   //-----------------------------
   // HP indication mixinghead 01:
   //-----------------------------
         A     "DB619_State_MPart".Recirculation[1].Lamp_HP."01";
         =     "DB123_MH_IO_Signals".MH[1].OUT.MH.H_HighPressure_MH;
   //-----
         A     "DB619_State_MPart".Recirculation[1].Highpressure;
         A(;
         L     "DB619_State_MPart".Recirculation[1].SWU_RC_HP;
         L     16#0000_0001;
         ==D;
         );
         =     "DB619_State_MPart".Recirculation[1].Indicator_HP."01";
         JCN   NoHP_MH01;
         L     1;
         T     "DB614_MH_State".MH_Status[1].State_HP;
   NoHP_MH01:NOP   0;
   //__________________________________________________________________
   //-----------------------------
   // HP indication mixinghead 02:
   //-----------------------------
         A     "DB619_State_MPart".Recirculation[1].Lamp_HP."02";
         =     "DB123_MH_IO_Signals".MH[2].OUT.MH.H_HighPressure_MH;
   //-----
         A     "DB619_State_MPart".Recirculation[1].Highpressure;
         A(;
         L     "DB619_State_MPart".Recirculation[1].SWU_RC_HP;
         L     16#0000_0002;
         ==D;
         );
         =     "DB619_State_MPart".Recirculation[1].Indicator_HP."02";
         JCN   NoHP_MH02;
         L     1;
         T     "DB614_MH_State".MH_Status[2].State_HP;
   NoHP_MH02:NOP   0;
   //___________________________________________________________________
   //-----------------------------
   // HP indication mixinghead 03:
   //-----------------------------
         A     "DB619_State_MPart".Recirculation[1].Lamp_HP."03";
         =     "DB123_MH_IO_Signals".MH[3].OUT.MH.H_HighPressure_MH;
   //-----
         A     "DB619_State_MPart".Recirculation[1].Highpressure;
         A(;
         L     "DB619_State_MPart".Recirculation[1].SWU_RC_HP;
         L     16#0000_0004;
         ==D;
         );
         =     "DB619_State_MPart".Recirculation[1].Indicator_HP."03";
         JCN   NoHP_MH03;
         L     1;
         T     "DB614_MH_State".MH_Status[3].State_HP;
   NoHP_MH03:NOP   0;
   //___________________________________________________________________
   //-----------------------------
   // HP indication mixinghead 04:
   //-----------------------------
         A     "DB619_State_MPart".Recirculation[1].Lamp_HP."04";
         =     "DB123_MH_IO_Signals".MH[4].OUT.MH.H_HighPressure_MH;
   //-----
         A     "DB619_State_MPart".Recirculation[1].Highpressure;
         A(;
         L     "DB619_State_MPart".Recirculation[1].SWU_RC_HP;
         L     16#0000_0008;
         ==D;
         );
         =     "DB619_State_MPart".Recirculation[1].Indicator_HP."04";
         JCN   NoHP_MH04;
         L     1;
         T     "DB614_MH_State".MH_Status[4].State_HP;
   NoHP_MH04:NOP   0;
   //___________________________________________________________________
   //-----------------------------
   // HP indication mixinghead 05:
   //-----------------------------
         A     "DB619_State_MPart".Recirculation[1].Lamp_HP."05";
         =     "DB123_MH_IO_Signals".MH[5].OUT.MH.H_HighPressure_MH;
   //-----
         A     "DB619_State_MPart".Recirculation[1].Highpressure;
         A(;
         L     "DB619_State_MPart".Recirculation[1].SWU_RC_HP;
         L     16#0000_0010;
         ==D;
         );
         =     "DB619_State_MPart".Recirculation[1].Indicator_HP."05";
         JCN   NoHP_MH05;
         L     1;
         T     "DB614_MH_State".MH_Status[5].State_HP;
   NoHP_MH05:NOP   0;
   //___________________________________________________________________
   //-----------------------------
   // HP indication mixinghead 06:
   //-----------------------------
         A     "DB619_State_MPart".Recirculation[1].Lamp_HP."06";
         =     "DB123_MH_IO_Signals".MH[6].OUT.MH.H_HighPressure_MH;
   //-----
         A     "DB619_State_MPart".Recirculation[1].Highpressure;
         A(;
         L     "DB619_State_MPart".Recirculation[1].SWU_RC_HP;
         L     16#0000_0020;
         ==D;
         );
         =     "DB619_State_MPart".Recirculation[1].Indicator_HP."06";
         JCN   NoHP_MH06;
         L     1;
         T     "DB614_MH_State".MH_Status[6].State_HP;
   NoHP_MH06:NOP   0;
   //___________________________________________________________________
   //-----------------------------
   // HP indication mixinghead 07:
   //-----------------------------
         A     "DB619_State_MPart".Recirculation[1].Lamp_HP."07";
         =     "DB123_MH_IO_Signals".MH[7].OUT.MH.H_HighPressure_MH;
   //-----
         A     "DB619_State_MPart".Recirculation[1].Highpressure;
         A(;
         L     "DB619_State_MPart".Recirculation[1].SWU_RC_HP;
         L     16#0000_0040;
         ==D;
         );
         =     "DB619_State_MPart".Recirculation[1].Indicator_HP."07";
         JCN   NoHP_MH07;
         L     1;
         T     "DB614_MH_State".MH_Status[7].State_HP;
   NoHP_MH07:NOP   0;
   //___________________________________________________________________
   //-----------------------------
   // HP indication mixinghead 08:
   //-----------------------------
         A     "DB619_State_MPart".Recirculation[1].Lamp_HP."08";
         =     "DB123_MH_IO_Signals".MH[8].OUT.MH.H_HighPressure_MH;
   //-----
         A     "DB619_State_MPart".Recirculation[1].Highpressure;
         A(;
         L     "DB619_State_MPart".Recirculation[1].SWU_RC_HP;
         L     16#0000_0080;
         ==D;
         );
         =     "DB619_State_MPart".Recirculation[1].Indicator_HP."08";
         JCN   NoHP_MH08;
         L     1;
         T     "DB614_MH_State".MH_Status[8].State_HP;
   NoHP_MH08:NOP   0;
   //___________________________________________________________________
   //-----------------------------
   // HP indication mixinghead 09:
   //-----------------------------
         A     "DB619_State_MPart".Recirculation[1].Lamp_HP."09";
         =     "DB123_MH_IO_Signals".MH[9].OUT.MH.H_HighPressure_MH;
   //-----
         A     "DB619_State_MPart".Recirculation[1].Highpressure;
         A(;
         L     "DB619_State_MPart".Recirculation[1].SWU_RC_HP;
         L     16#0000_0100;
         ==D;
         );
         =     "DB619_State_MPart".Recirculation[1].Indicator_HP."09";
         JCN   NoHP_MH09;
         L     1;
         T     "DB614_MH_State".MH_Status[9].State_HP;
   NoHP_MH09:NOP   0;
   //___________________________________________________________________
   //-----------------------------
   // HP indication mixinghead 10:
   //-----------------------------
         A     "DB619_State_MPart".Recirculation[1].Lamp_HP."10";
         =     "DB123_MH_IO_Signals".MH[10].OUT.MH.H_HighPressure_MH;
   //-----
         A     "DB619_State_MPart".Recirculation[1].Highpressure;
         A(;
         L     "DB619_State_MPart".Recirculation[1].SWU_RC_HP;
         L     16#0000_0200;
         ==D;
         );
         =     "DB619_State_MPart".Recirculation[1].Indicator_HP."10";
         JCN   NoHP_MH10;
         L     1;
         T     "DB614_MH_State".MH_Status[10].State_HP;
   NoHP_MH10:NOP   0;
   //___________________________________________________________________
   //-----------------------------
   // HP indication mixinghead 11:
   //-----------------------------
         A     "DB619_State_MPart".Recirculation[1].Lamp_HP."11";
         =     "DB123_MH_IO_Signals".MH[11].OUT.MH.H_HighPressure_MH;
   //-----
         A     "DB619_State_MPart".Recirculation[1].Highpressure;
         A(;
         L     "DB619_State_MPart".Recirculation[1].SWU_RC_HP;
         L     16#0000_0400;
         ==D;
         );
         =     "DB619_State_MPart".Recirculation[1].Indicator_HP."11";
         JCN   NoHP_MH11;
         L     1;
         T     "DB614_MH_State".MH_Status[11].State_HP;
   NoHP_MH11:NOP   0;
   //___________________________________________________________________
   //-----------------------------
   // HP indication mixinghead 12:
   //-----------------------------
         A     "DB619_State_MPart".Recirculation[1].Lamp_HP."12";
         =     "DB123_MH_IO_Signals".MH[12].OUT.MH.H_HighPressure_MH;
   //-----
         A     "DB619_State_MPart".Recirculation[1].Highpressure;
         A(;
         L     "DB619_State_MPart".Recirculation[1].SWU_RC_HP;
         L     16#0000_0800;
         ==D;
         );
         =     "DB619_State_MPart".Recirculation[1].Indicator_HP."12";
         JCN   NoHP_MH12;
         L     1;
         T     "DB614_MH_State".MH_Status[12].State_HP;
   NoHP_MH12:NOP   0;
   //___________________________________________________________________
   //
END_REGION

REGION Network 13: Activate valve of low pressure cycle
         O     "DB619_State_MPart".Machine[1].Metering."01";
         O     "DB619_State_MPart".Machine[1].Metering."02";
         O     "DB619_State_MPart".Machine[1].Metering."03";
         O     "DB619_State_MPart".Machine[1].Metering."04";
         A     "DB619_State_MPart".Machine[1].HydStartUp_finished;
         L     "DB700_Machine".Machine[1].LP_Valve_switchOFF_Delay;
         SF    "TM_Kreislauf_ND_M1";
   //
         A(;
         O     "DB619_State_MPart".Recirculation[1].Lowpressure;
         ON    "DB619_State_MPart".Recirculation[1].Is_active;
         A     "TM_Kreislauf_ND_M1";
         );
         AN    "DB619_State_MPart".Cycle[1].running;
   //      NOT                        // <- Depending of the low pressure valve
         =     #Temp_HF_LP_circ;
   //
         A     "DB619_State_MPart".SWU[1].Open_SWU_allone."01";
         A     #Temp_HF_LP_circ;
         =     "DB123_MH_IO_Signals".MH[1].OUT.MH.V_LowPressure_Circ_MH;
   //
         A     "DB619_State_MPart".SWU[1].Open_SWU_allone."02";
         A     #Temp_HF_LP_circ;
         =     "DB123_MH_IO_Signals".MH[2].OUT.MH.V_LowPressure_Circ_MH;
   //
         A     "DB619_State_MPart".SWU[1].Open_SWU_allone."03";
         A     #Temp_HF_LP_circ;
         =     "DB123_MH_IO_Signals".MH[3].OUT.MH.V_LowPressure_Circ_MH;
   //
         A     "DB619_State_MPart".SWU[1].Open_SWU_allone."04";
         A     #Temp_HF_LP_circ;
         =     "DB123_MH_IO_Signals".MH[4].OUT.MH.V_LowPressure_Circ_MH;
   //
         A     "DB619_State_MPart".SWU[1].Open_SWU_allone."05";
         A     #Temp_HF_LP_circ;
         =     "DB123_MH_IO_Signals".MH[5].OUT.MH.V_LowPressure_Circ_MH;
   //
         A     "DB619_State_MPart".SWU[1].Open_SWU_allone."06";
         A     #Temp_HF_LP_circ;
         =     "DB123_MH_IO_Signals".MH[6].OUT.MH.V_LowPressure_Circ_MH;
   //
         A     "DB619_State_MPart".SWU[1].Open_SWU_allone."07";
         A     #Temp_HF_LP_circ;
         =     "DB123_MH_IO_Signals".MH[7].OUT.MH.V_LowPressure_Circ_MH;
   //
         A     "DB619_State_MPart".SWU[1].Open_SWU_allone."08";
         A     #Temp_HF_LP_circ;
         =     "DB123_MH_IO_Signals".MH[8].OUT.MH.V_LowPressure_Circ_MH;
   //
         A     "DB619_State_MPart".SWU[1].Open_SWU_allone."09";
         A     #Temp_HF_LP_circ;
         =     "DB123_MH_IO_Signals".MH[9].OUT.MH.V_LowPressure_Circ_MH;
   //
         A     "DB619_State_MPart".SWU[1].Open_SWU_allone."10";
         A     #Temp_HF_LP_circ;
         =     "DB123_MH_IO_Signals".MH[10].OUT.MH.V_LowPressure_Circ_MH;
   //
         A     "DB619_State_MPart".SWU[1].Open_SWU_allone."11";
         A     #Temp_HF_LP_circ;
         =     "DB123_MH_IO_Signals".MH[11].OUT.MH.V_LowPressure_Circ_MH;
   //
         A     "DB619_State_MPart".SWU[1].Open_SWU_allone."12";
         A     #Temp_HF_LP_circ;
         =     "DB123_MH_IO_Signals".MH[12].OUT.MH.V_LowPressure_Circ_MH;
   //
END_REGION
END_FUNCTION_BLOCK

FUNCTION_BLOCK "FB012_MH_Hydraulic_M1"   // FB12, STL
TITLE = Hydraulics and elapsed hour meter
{ S7_Optimized_Access := 'FALSE' }
AUTHOR : KT242
VERSION : 0.1
// Hydraulic and elapsed hour meter
   VAR_TEMP
      Temp_P_top_MH_Hydr : Bool;
      Temp_L_Oil_Hydraulic : Bool;
      Temp_C_Oil : Bool;
      Temp_MachineHourCounter : Bool;
      Temp_M_Hydr_PowerSupply : Bool;
      Temp_M_Hydr_Star : Bool;
      Temp_M_Hydr_Delta : Bool;
      Temp_V_Oel_Cooling : Bool;
      Temp_P_Max_Hydraulic : Bool;
      Temp_Hydraulic_active : Bool;
      Temp_PausTime : Bool;
      Temp_PhydraulicOK : Bool;
      RTM_NR_0 : Byte;
      RET_VAL_0 : Int;
      ExternalFault : Bool;
      RTM_NR : Byte;
      RTM_MODE : Byte;
      RetValSFC : Int;
      _Accu1Safe : DInt;
      _Accu2Safe : DInt;
      Migra_NR : Rtm;
   END_VAR
BEGIN

REGION Network 1: Mixinghead hydraulic
   //-----
         O(;
         ON    "DB721_MH_Hydraulic".Option[1].With2PSwitch;
         ON    "DB619_State_MPart".Cycle[1].SelectHydForShot;
         A     "P_MK_Hydr";
         );
         O(;
         A     "DB721_MH_Hydraulic".Option[1].With2PSwitch;
         A     "DB619_State_MPart".Cycle[1].SelectHydForShot;
         A     "P_2_MK_Hydr";
         );
         =     #Temp_PhydraulicOK;
   //-----
         A     #Temp_PhydraulicOK;
         L     "DB721_MH_Hydraulic".MH_Hyd[1].Hyd_PressureSwitch;
         SD    "TM_P_oben_MK_Hyd_M1";
         AN    "TM_P_oben_MK_Hyd_M1";
         =     #Temp_P_top_MH_Hydr;  // für RS- Maschinen

   //-----
         A(;
         ON    "DB613_Komponent_State".MeteringPump[1].Selection_Feedingpump;
         ON    "DB753_MeteringPump".Pump[1].WithFeedPump;
         ON    "DB753_MeteringPump".Pump[1].Pump_Active;
         );
         A(;
         ON    "DB613_Komponent_State".MeteringPump[2].Selection_Feedingpump;
         ON    "DB753_MeteringPump".Pump[2].WithFeedPump;
         ON    "DB753_MeteringPump".Pump[2].Pump_Active;
         );
         A     "DB619_State_MPart".Recirculation[1].Pausetime;
         =     #Temp_PausTime;
   //-----
         CALL  "FC021_MH_Hydraulic"
         ( IN_MotorProtection       := "F_MK_Hydr",
           IN_Min_Level             := "L_Min_Oel_MK_Hydr",
           IN_C_OilCooling          := "C_Cooling_Hydr",
           IN_C_Max                 := "C_Max_Oel_MK_Hydr",
           IN_F_Filter_FeedLine     := "F_Fil_MK_Hydr_VL",
           IN_F_Filter_ReturnLine   := TRUE,
           IN_OPMode_Automatic      := "DB619_State_MPart".Operationmode[1].Auto,
           IN_OPMode_Manual         := "DB619_State_MPart".Operationmode[1].Manual,
           IN_PauseTime             := #Temp_PausTime,  // "DB619_State_MPart".Recirculation[1].Pausetime
           IN_Pos_of_Pause_ok       := "DB619_State_MPart".CylinderManager[1].Pos_Weekends_Pause,
           IN_Fault_from_Extern     := FALSE,
           IN_P_lowerlimit          := #Temp_PhydraulicOK,
           IN_P_upperLimit          := #Temp_P_top_MH_Hydr,
           IN_Option2SetPoints      := "DB721_MH_Hydraulic".Option[1].With2PSwitch,
           IN_PRequestCycle         := "DB619_State_MPart".Cycle[1].SelectHydForShot,
           IN_KK_Manager_active     := FALSE,
           IN_ShotStroke_by_Piston  := FALSE,
           IN_Reset_fault_Fkt       := "DB009_Faults".Faults_Reset_FKT_M1,
           IN_Temperatur_Timer      := "TM_MK_Hyd_Temp_M1",
           IN_Filter_Timer          := "TM_MK_Hyd_Filter_M1",
           IN_Hydraulictimer        := "TM_MK_Hyd_M1",
           IN_Star_Delta_Timer      := S5T#1S,
           IN_Delay_FilterError     := "DB721_MH_Hydraulic".MH_Hyd[1].Hyd_Filter_supervision,
           IN_P_BuildUpTime         := "DB721_MH_Hydraulic".MH_Hyd[1].Hyd_P_Startup,
           IN_P_OperationTime       := "DB721_MH_Hydraulic".MH_Hyd[1].Hyd_P_Supervision,
           IN_P_ClPistonTime        := "DB721_MH_Hydraulic".MH_Hyd[1].Hyd_CP_Time,
           IN_SwitchOffTime         := "DB721_MH_Hydraulic".MH_Hyd[1].Hyd_SwitchOFFDelay,
           IN_SwitchOFFTimer        := "TM_SwitchOffHydMH_M1",
           OUT_Hydraulic_active     := #Temp_Hydraulic_active,
           OUT_PressureValve        := "V_P_builtup_MH_Hydr_M1",
           OUT_Motor_MainsContactor := "M_MH_Hydr_Net_M1",
           OUT_Motor_Star           := #Temp_M_Hydr_Star,
           OUT_Motor_Delta          := #Temp_M_Hydr_Delta,
           OUT_V_OilCooling         := "V_Cooling_Hydr",
           IO_Status                := "DB611_Hydraulic_State".MH_Hydraulic[1],
           IO_Fault                 := "DB821_Error_Hydraulic".MH_Hydraulic[1],
           IO_NewFault              := "DB009_Faults".Faultschanging_M1,
           IO_FaultLevel_1          := "DB009_Faults".Faults_FKT_Grp_1_M1,
           IO_FaultLevel_2          := "DB009_Faults".Faults_FKT_Grp_2_M1,
           IO_FaultLevel_3          := "DB009_Faults".Faults_FKT_Grp_3_M1
         );
   //
         A     "DB611_Hydraulic_State".MH_Hydraulic[1].Request_from_CP;
         L     S5T#1M;
         SD    "TM_Hydraulik_RK_Druck";
         A     "TM_Hydraulik_RK_Druck";
         R     "DB611_Hydraulic_State".MH_Hydraulic[1].Request_from_CP;
   //
END_REGION

REGION Network 2: Hydraulic start up finished
         A     "DB611_Hydraulic_State".MH_Hydraulic[1].MH_Hyd_OK;
         =     "DB619_State_MPart".Machine[1].HydStartUp_finished;
END_REGION

REGION Network 3: Machine operation hour counter
         L     0;
         T     #RTM_NR;
   //
         L     16#01;  // Mode 1: Start counter
         A     "DB619_State_MPart".Machine[1].HydStartUp_finished;
         AN    "M_RTM0Running";
         JC    mode;

         L     16#02;  // Mode 2: Stop counter
         AN    "DB619_State_MPart".Machine[1].HydStartUp_finished;
         A     "M_RTM0Running";
         JC    mode;
         L     16#00;  // Mode 0: Read counter
   mode: T     #RTM_MODE;

         T     #_Accu1Safe;
         TAK;
         T     #_Accu2Safe;
         L     #RTM_NR;
         T     #Migra_NR;
         CALL  RTM
         ( NR      := #Migra_NR,
           MODE    := #RTM_MODE,
           PV      := 0,
           RET_VAL := #RetValSFC,
           CQ      := "M_RTM0Running",
           CV      := "DB611_Hydraulic_State".MH_Hydraulic[1].HourCounter
         );
         L     #_Accu2Safe;
         L     #_Accu1Safe;
END_REGION
END_FUNCTION_BLOCK

FUNCTION_BLOCK "FB014_MH_SWU_M1"   // FB14, STL
TITLE = Activation of mixingheads and switch over units (SWU)
{ S7_Optimized_Access := 'FALSE' }
AUTHOR : KT242
VERSION : 0.1
   VAR_TEMP
      Dummy_Schusszaehler : Bool;
      Temp_OperationMode : Bool;
      Nullbyte : Byte;
      RetValSFC : Int;
      SWU_DWORD : DWord;
      TempMask : Struct
         ForceNozzle_1 : Bool;
         ForceNozzle_2 : Bool;
         ForceNozzle_3 : Bool;
         ForceNozzle_4 : Bool;
         ForceNozzle_5 : Bool;
         ForceNozzle_6 : Bool;
         ForceNozzle_7 : Bool;
         ForceNozzle_8 : Bool;
         EnableNozzle_1 : Bool;
         EnableNozzle_2 : Bool;
         EnableNozzle_3 : Bool;
         EnableNozzle_4 : Bool;
         EnableNozzle_5 : Bool;
         EnableNozzle_6 : Bool;
         EnableNozzle_7 : Bool;
         EnableNozzle_8 : Bool;
      END_STRUCT;
      TempNozzleShotConnection : Array[1..8] of Bool;
      TempNozzleCirc : Array[1..8] of Bool;
      TempNozzleShotMH : Array[1..8] of Bool;
      SwitchOff : Word;
      SwitchOn : Word;
   END_VAR
BEGIN

REGION Network 1: Release to switch over to different mixingheads
   // Set SWU  release of 32 mixingheads to zero
         L     0;
         T     #Nullbyte;
         CALL  FILL
         ( BVAL    := #Nullbyte,
           RET_VAL := #RetValSFC,
           BLK     := "DB619_State_MPart".SWU[1].SWU_released
         );
   //__________________________________________________________________
   // For mixinghead 01:
   //
         L     "DB704_MH_Value".Mixinghead[1].MachineNumber;
         L     1;
         ==D;
         JCN   Nsel_MH01;
   //-
         L     "DB790_PlantParameter".AmountMH;
         L     1;
         ==D;
         O     "DB123_MH_IO_Signals".MH[1].IN.MH_Release_SWU;
         =     "DB619_State_MPart".SWU[1].SWU_released."01";
         =     "DB614_MH_State".MH_Status[1].SWU_released;
   Nsel_MH01:NOP   0;
   //__________________________________________________________________
   // For mixinghead 02:
         L     "DB704_MH_Value".Mixinghead[2].MachineNumber;
         L     1;
         ==D;
         JCN   Nsel_MH02;
   //-
         L     "DB790_PlantParameter".AmountMH;
         L     2;
         <D;
         JC    swue;
         A     "DB123_MH_IO_Signals".MH[2].IN.MH_Release_SWU;
         =     "DB619_State_MPart".SWU[1].SWU_released."02";
         =     "DB614_MH_State".MH_Status[2].SWU_released;
   Nsel_MH02:NOP   0;
   //__________________________________________________________________
   // For mixinghead 03:
         L     "DB704_MH_Value".Mixinghead[3].MachineNumber;
         L     1;
         ==D;
         JCN   Nsel_MH03;
   //-
         L     "DB790_PlantParameter".AmountMH;
         L     3;
         <D;
         JC    swue;
         A     "DB123_MH_IO_Signals".MH[3].IN.MH_Release_SWU;
         =     "DB619_State_MPart".SWU[1].SWU_released."03";
         =     "DB614_MH_State".MH_Status[3].SWU_released;
   Nsel_MH03:NOP   0;
   //__________________________________________________________________
   // For mixinghead 04:
         L     "DB704_MH_Value".Mixinghead[4].MachineNumber;
         L     1;
         ==D;
         JCN   Nsel_MH04;
   //-
         L     "DB790_PlantParameter".AmountMH;
         L     4;
         <D;
         JC    swue;
         A     "DB123_MH_IO_Signals".MH[4].IN.MH_Release_SWU;
         =     "DB619_State_MPart".SWU[1].SWU_released."04";
         =     "DB614_MH_State".MH_Status[4].SWU_released;
   Nsel_MH04:NOP   0;
   //__________________________________________________________________
   // For mixinghead 05:
         L     "DB704_MH_Value".Mixinghead[5].MachineNumber;
         L     1;
         ==D;
         JCN   Nsel_MH05;
   //-
         L     "DB790_PlantParameter".AmountMH;
         L     5;
         <D;
         JC    swue;
         A     "DB123_MH_IO_Signals".MH[5].IN.MH_Release_SWU;
         =     "DB619_State_MPart".SWU[1].SWU_released."05";
         =     "DB614_MH_State".MH_Status[5].SWU_released;
   Nsel_MH05:NOP   0;
   //__________________________________________________________________
   // For mixinghead 06:
         L     "DB704_MH_Value".Mixinghead[6].MachineNumber;
         L     1;
         ==D;
         JCN   Nsel_MH06;
   //-
         L     "DB790_PlantParameter".AmountMH;
         L     6;
         <D;
         JC    swue;
         A     "DB123_MH_IO_Signals".MH[6].IN.MH_Release_SWU;
         =     "DB619_State_MPart".SWU[1].SWU_released."06";
         =     "DB614_MH_State".MH_Status[6].SWU_released;
   Nsel_MH06:NOP   0;
   //__________________________________________________________________
   // For mixinghead 07:
         L     "DB704_MH_Value".Mixinghead[7].MachineNumber;
         L     1;
         ==D;
         JCN   Nsel_MH07;
   //-
         L     "DB790_PlantParameter".AmountMH;
         L     7;
         <D;
         JC    swue;
         A     "DB123_MH_IO_Signals".MH[7].IN.MH_Release_SWU;
         =     "DB619_State_MPart".SWU[1].SWU_released."07";
         =     "DB614_MH_State".MH_Status[7].SWU_released;
   Nsel_MH07:NOP   0;
   //__________________________________________________________________
   // For mixinghead 08:
         L     "DB704_MH_Value".Mixinghead[8].MachineNumber;
         L     1;
         ==D;
         JCN   Nsel_MH08;
   //-
         L     "DB790_PlantParameter".AmountMH;
         L     8;
         <D;
         JC    swue;
         A     "DB123_MH_IO_Signals".MH[8].IN.MH_Release_SWU;
         =     "DB619_State_MPart".SWU[1].SWU_released."08";
         =     "DB614_MH_State".MH_Status[8].SWU_released;
   Nsel_MH08:NOP   0;
   //__________________________________________________________________
   // For mixinghead 09:
         L     "DB704_MH_Value".Mixinghead[9].MachineNumber;
         L     1;
         ==D;
         JCN   Nsel_MH09;
   //-
         L     "DB790_PlantParameter".AmountMH;
         L     9;
         <D;
         JC    swue;
         A     "DB123_MH_IO_Signals".MH[9].IN.MH_Release_SWU;
         =     "DB619_State_MPart".SWU[1].SWU_released."09";
         =     "DB614_MH_State".MH_Status[9].SWU_released;
   Nsel_MH09:NOP   0;
   //__________________________________________________________________
   // For mixinghead 10:
         L     "DB704_MH_Value".Mixinghead[10].MachineNumber;
         L     1;
         ==D;
         JCN   Nsel_MH10;
   //-
         L     "DB790_PlantParameter".AmountMH;
         L     10;
         <D;
         JC    swue;
         A     "DB123_MH_IO_Signals".MH[10].IN.MH_Release_SWU;
         =     "DB619_State_MPart".SWU[1].SWU_released."10";
         =     "DB614_MH_State".MH_Status[10].SWU_released;
   Nsel_MH10:NOP   0;
   //__________________________________________________________________
   //
   swue: NOP   0;
   //------------------------------------------------------------------
   //  Get info about MH at machine
   //------------------------------------------------------------------
         CALL  BLKMOV
         ( SRCBLK  := "DB619_State_MPart".SWU[1].SWU_released,
           RET_VAL := #RetValSFC,
           DSTBLK  := "DB619_State_MPart".MH_at_Machine[1]
         );

   // "DB700_Machine".Machine[1].MH_at_Machine wird nur noch im FB1930 "GetToolShotValues" verwendet
   // sollte auch anders gelöst werden!! vdG 20140322
         CALL  BLKMOV
         ( SRCBLK  := "DB619_State_MPart".MH_at_Machine[1],
           RET_VAL := #RetValSFC,
           DSTBLK  := "DB700_Machine".Machine[1].MH_at_Machine
         );
END_REGION

REGION Network 2: Selection of SWU 1..32 (SWU -> Switch over unit)
         CALL  "FC041_SwitchOverUnit"
         ( IN_select_piston         := "DB619_State_MPart".CylinderManager[1].Block_is_active,
           IN_filling_piston        := "DB619_State_MPart".CylinderManager[1].Selection_Filling,
           IN_OperationMode_valid   := "DB619_State_MPart".Operationmode[1].valid,
           IN_AcknoldgeFaults       := "DB009_Faults".Faults_Reset_FKT_M1,
           IN_cycle_running         := "DB619_State_MPart".Cycle[1].running,
           IN_PistonService         := "DB619_State_MPart".Operationmode[1].Cylinderservice,
           IN_Circulation_active    := "DB619_State_MPart".Recirculation[1].Is_active,
           IN_Circulation_HP_active := "DB619_State_MPart".Recirculation[1].HP_is_active,
           IN_MH_No_at_FoamingCycle := "DB619_State_MPart".ShotMa[1].ShotData.MH_No,
           IN_MH_No_at_HP_Cycle     := "DB619_State_MPart".Recirculation[1].SWU_RC_HP,
           IN_StokeCounter          := "Z_HubzaehlerM1",
           IN_Amount_Strokes        := "DB700_Machine".Machine[1].StrokeCounter_KK,
           IN_FlushingTimer         := "TM_USE_Taktzeit_M1",
           IN_SWU_FlushingTime      := "DB700_Machine".Machine[1].SWU_Intervalltime,
           IN_SwitchOverTimer       := "TM_USE_Umschaltzeit_M1",
           IN_SwitchOffTime         := S5T#5S,
           IN_SwitchOverTime        := S5T#1S,
           IO_Status                := "DB619_State_MPart".SWU[1],
           IO_Fault                 := "DB829_Error_Machine".SWU[1],
           IO_NewFault              := "DB009_Faults".Faultschanging_M1,
           IO_FaultLevel_1          := "DB009_Faults".Faults_FKT_Grp_1_M1,
           IO_FaultLevel_2          := "DB009_Faults".Faults_FKT_Grp_2_M1,
           IO_FaultLevel_3          := "DB009_Faults".Faults_FKT_Grp_3_M1
         );
   //
END_REGION

REGION Network 3: Open SWU
   //__________________________________________________________________
   // SWU mixinghead 01:
   //
         L     "DB704_MH_Value".Mixinghead[1].MachineNumber;
         L     1;
         <=D;
         JCN   NSWU_MH01;
         A     "DB619_State_MPart".SWU[1].Open_SWU."01";
         =     "DB123_MH_IO_Signals".MH[1].OUT.MH.V_SWU_MH;
   NSWU_MH01:NOP   0;
   //__________________________________________________________________
   // SWU mixinghead 02:
         L     "DB704_MH_Value".Mixinghead[2].MachineNumber;
         L     1;
         <=D;
         JCN   NSWU_MH02;
         A     "DB619_State_MPart".SWU[1].Open_SWU."02";
         =     "DB123_MH_IO_Signals".MH[2].OUT.MH.V_SWU_MH;
   NSWU_MH02:NOP   0;
   //__________________________________________________________________
   // SWU mixinghead 03:
   //
         L     "DB704_MH_Value".Mixinghead[3].MachineNumber;
         L     1;
         <=D;
         JCN   NSWU_MH03;
         A     "DB619_State_MPart".SWU[1].Open_SWU."03";
         =     "DB123_MH_IO_Signals".MH[3].OUT.MH.V_SWU_MH;
   NSWU_MH03:NOP   0;
   //__________________________________________________________________
   // SWU mixinghead 04:
   //
         L     "DB704_MH_Value".Mixinghead[4].MachineNumber;
         L     1;
         <=D;
         JCN   NSWU_MH04;
         A     "DB619_State_MPart".SWU[1].Open_SWU."04";
         =     "DB123_MH_IO_Signals".MH[4].OUT.MH.V_SWU_MH;
   NSWU_MH04:NOP   0;
   //__________________________________________________________________
   // SWU mixinghead 05:
   //
         L     "DB704_MH_Value".Mixinghead[5].MachineNumber;
         L     1;
         <=D;
         JCN   NSWU_MH05;
         A     "DB619_State_MPart".SWU[1].Open_SWU."05";
         =     "DB123_MH_IO_Signals".MH[5].OUT.MH.V_SWU_MH;
   NSWU_MH05:NOP   0;
   //__________________________________________________________________
   // SWU mixinghead 06:
   //
         L     "DB704_MH_Value".Mixinghead[6].MachineNumber;
         L     1;
         <=D;
         JCN   NSWU_MH06;
         A     "DB619_State_MPart".SWU[1].Open_SWU."06";
         =     "DB123_MH_IO_Signals".MH[6].OUT.MH.V_SWU_MH;
   NSWU_MH06:NOP   0;
   //__________________________________________________________________
   // SWU mixinghead 07:
   //
         L     "DB704_MH_Value".Mixinghead[7].MachineNumber;
         L     1;
         <=D;
         JCN   NSWU_MH07;
         A     "DB619_State_MPart".SWU[1].Open_SWU."07";
         =     "DB123_MH_IO_Signals".MH[7].OUT.MH.V_SWU_MH;
   NSWU_MH07:NOP   0;
   //__________________________________________________________________
   // SWU mixinghead 08:
   //
         L     "DB704_MH_Value".Mixinghead[8].MachineNumber;
         L     1;
         <=D;
         JCN   NSWU_MH08;
         A     "DB619_State_MPart".SWU[1].Open_SWU."08";
         =     "DB123_MH_IO_Signals".MH[8].OUT.MH.V_SWU_MH;
   NSWU_MH08:NOP   0;
   //__________________________________________________________________
   // SWU mixinghead 09:
   //
         L     "DB704_MH_Value".Mixinghead[9].MachineNumber;
         L     1;
         <=D;
         JCN   NSWU_MH09;
         A     "DB619_State_MPart".SWU[1].Open_SWU."09";
         =     "DB123_MH_IO_Signals".MH[9].OUT.MH.V_SWU_MH;
   NSWU_MH09:NOP   0;
   //__________________________________________________________________
   // SWU mixinghead 10:
   //
         L     "DB704_MH_Value".Mixinghead[10].MachineNumber;
         L     1;
         <=D;
         JCN   NSWU_MH10;
         A     "DB619_State_MPart".SWU[1].Open_SWU."10";
         =     "DB123_MH_IO_Signals".MH[10].OUT.MH.V_SWU_MH;
   NSWU_MH10:NOP   0;
   //__________________________________________________________________
   //
END_REGION

REGION Network 4: Releases to open mixinghead
   //__________________________________________________________________
   // Releases Mixinghead 01:
   //
         A(;
         A     "DB614_MH_State".MH_Status[1].OpenMHEnableExtern;
         A     "DB704_MH_Value".Mixinghead[1].Conf_IntWithRobot;
         O;
         AN    "DB704_MH_Value".Mixinghead[1].Conf_IntWithRobot;
         A     "DB005_RS<->Extern".MC_Interface[1].Data_from_MC.Shot_release;
         A     "DB110_Interf_Program_M1".Status_IF[1].IF_is_on_1_Position;
         );
         A     "DB123_MH_IO_Signals".MH[1].IN.MH_Auto_Mode;
         O(;
         A     "DB123_MH_IO_Signals".MH[1].IN.MH_Manual_Mode;
         A     "DB110_Interf_Program_M1".Status_IF[1].IF_is_on_1_Position;
         );
         O     "DB619_State_MPart".Operationmode[1].Test;
         A(;
         O     "DB619_State_MPart".CylinderManager[1].Shothub;
         ON    "DB619_State_MPart".CylinderManager[1].Block_is_active;
         );
         =     "DB619_State_MPart".Mixinghead[1].Release_MH."01";
   //__________________________________________________________________
   // Releases Mixinghead 02:
   //
         A     "DB005_RS<->Extern".MC_Interface[2].Data_from_MC.Shot_release;
         A     "DB123_MH_IO_Signals".MH[2].IN.MH_Auto_Mode;
         O     "DB123_MH_IO_Signals".MH[2].IN.MH_Manual_Mode;
         A     "DB110_Interf_Program_M1".Status_IF[2].IF_is_on_1_Position;
         O     "DB619_State_MPart".Operationmode[1].Test;
         A(;
         O     "DB619_State_MPart".CylinderManager[1].Shothub;
         ON    "DB619_State_MPart".CylinderManager[1].Block_is_active;
         );
         AN    "DB824_Error_MH_CP".MH_Control[2].FLT_ShotStopped;
         =     "DB619_State_MPart".Mixinghead[1].Release_MH."02";
   //__________________________________________________________________
   // Releases Mixinghead 03:
   //
         A     "DB005_RS<->Extern".MC_Interface[3].Data_from_MC.Shot_release;
         A     "DB123_MH_IO_Signals".MH[3].IN.MH_Auto_Mode;
         O     "DB123_MH_IO_Signals".MH[3].IN.MH_Manual_Mode;
         A     "DB110_Interf_Program_M1".Status_IF[3].IF_is_on_1_Position;
         O     "DB619_State_MPart".Operationmode[1].Test;
         A(;
         O     "DB619_State_MPart".CylinderManager[1].Shothub;
         ON    "DB619_State_MPart".CylinderManager[1].Block_is_active;
         );
         =     "DB619_State_MPart".Mixinghead[1].Release_MH."03";
   //__________________________________________________________________
   // Releases Mixinghead 04:
   //
         A     "DB005_RS<->Extern".MC_Interface[4].Data_from_MC.Shot_release;
         A     "DB123_MH_IO_Signals".MH[4].IN.MH_Auto_Mode;
         O     "DB123_MH_IO_Signals".MH[4].IN.MH_Manual_Mode;
         A     "DB110_Interf_Program_M1".Status_IF[4].IF_is_on_1_Position;
         O     "DB619_State_MPart".Operationmode[1].Test;
         A(;
         O     "DB619_State_MPart".CylinderManager[1].Shothub;
         ON    "DB619_State_MPart".CylinderManager[1].Block_is_active;
         );
         =     "DB619_State_MPart".Mixinghead[1].Release_MH."04";
   //__________________________________________________________________
   // Releases Mixinghead 05:
   //
         A     "DB005_RS<->Extern".MC_Interface[5].Data_from_MC.Shot_release;
         A     "DB123_MH_IO_Signals".MH[5].IN.MH_Auto_Mode;
         O     "DB123_MH_IO_Signals".MH[5].IN.MH_Manual_Mode;
         A     "DB110_Interf_Program_M1".Status_IF[5].IF_is_on_1_Position;
         O     "DB619_State_MPart".Operationmode[1].Test;
         A(;
         O     "DB619_State_MPart".CylinderManager[1].Shothub;
         ON    "DB619_State_MPart".CylinderManager[1].Block_is_active;
         );
         =     "DB619_State_MPart".Mixinghead[1].Release_MH."05";
   //__________________________________________________________________
   // Releases Mixinghead 06:
   //
         A     "DB005_RS<->Extern".MC_Interface[6].Data_from_MC.Shot_release;
         A     "DB123_MH_IO_Signals".MH[6].IN.MH_Auto_Mode;
         O     "DB123_MH_IO_Signals".MH[6].IN.MH_Manual_Mode;
         A     "DB110_Interf_Program_M1".Status_IF[6].IF_is_on_1_Position;
         O     "DB619_State_MPart".Operationmode[1].Test;
         A(;
         O     "DB619_State_MPart".CylinderManager[1].Shothub;
         ON    "DB619_State_MPart".CylinderManager[1].Block_is_active;
         );
         =     "DB619_State_MPart".Mixinghead[1].Release_MH."06";
   //__________________________________________________________________
   // Releases Mixinghead 07:
   //
         A     "DB005_RS<->Extern".MC_Interface[7].Data_from_MC.Shot_release;
         A     "DB123_MH_IO_Signals".MH[7].IN.MH_Auto_Mode;
         O     "DB123_MH_IO_Signals".MH[7].IN.MH_Manual_Mode;
         A     "DB110_Interf_Program_M1".Status_IF[7].IF_is_on_1_Position;
         O     "DB619_State_MPart".Operationmode[1].Test;
         A(;
         O     "DB619_State_MPart".CylinderManager[1].Shothub;
         ON    "DB619_State_MPart".CylinderManager[1].Block_is_active;
         );
         =     "DB619_State_MPart".Mixinghead[1].Release_MH."07";
   //__________________________________________________________________
   // Releases Mixinghead 08:
   //
         A     "DB005_RS<->Extern".MC_Interface[8].Data_from_MC.Shot_release;
         A     "DB123_MH_IO_Signals".MH[8].IN.MH_Auto_Mode;
         O     "DB123_MH_IO_Signals".MH[8].IN.MH_Manual_Mode;
         A     "DB110_Interf_Program_M1".Status_IF[8].IF_is_on_1_Position;
         O     "DB619_State_MPart".Operationmode[1].Test;
         A(;
         O     "DB619_State_MPart".CylinderManager[1].Shothub;
         ON    "DB619_State_MPart".CylinderManager[1].Block_is_active;
         );
         =     "DB619_State_MPart".Mixinghead[1].Release_MH."08";
   //__________________________________________________________________
   // Releases Mixinghead 09:
   //
         A     "DB123_MH_IO_Signals".MH[9].IN.MH_Releas_Foaming_MC;
         A     "DB123_MH_IO_Signals".MH[9].IN.MH_Auto_Mode;
         O     "DB123_MH_IO_Signals".MH[9].IN.MH_Manual_Mode;
         A     "DB110_Interf_Program_M1".Status_IF[9].IF_is_on_1_Position;
         O     "DB619_State_MPart".Operationmode[1].Test;
         A(;
         O     "DB619_State_MPart".CylinderManager[1].Shothub;
         ON    "DB619_State_MPart".CylinderManager[1].Block_is_active;
         );
         =     "DB619_State_MPart".Mixinghead[1].Release_MH."09";
   //__________________________________________________________________
   // Releases Mixinghead 10:
   //
         A     "DB005_RS<->Extern".MC_Interface[10].Data_from_MC.Shot_release;
         A     "DB123_MH_IO_Signals".MH[10].IN.MH_Auto_Mode;
         O     "DB123_MH_IO_Signals".MH[10].IN.MH_Manual_Mode;
         A     "DB110_Interf_Program_M1".Status_IF[10].IF_is_on_1_Position;
         O     "DB619_State_MPart".Operationmode[1].Test;
         A(;
         O     "DB619_State_MPart".CylinderManager[1].Shothub;
         ON    "DB619_State_MPart".CylinderManager[1].Block_is_active;
         );
         =     "DB619_State_MPart".Mixinghead[1].Release_MH."10";
   //__________________________________________________________________
   //
END_REGION

REGION Network 5: Selection of mixingheads 1..32
   //-----
         A     "DB619_State_MPart".Operationmode[1].Operation;
         AN    "DB619_State_MPart".ShotMa[1].ShotData.ShotDisabled;
         =     #Temp_OperationMode;
   //-----
         CALL  "FC042_MixingHead"
         ( IN_SWU_openValve        := "DB619_State_MPart".SWU[1].Target_SWU,
           IN_OPMode_Automatic     := "DB619_State_MPart".Operationmode[1].Auto,
           IN_OPMode_Production    := #Temp_OperationMode,
           IN_OPMode_Test          := "DB619_State_MPart".Operationmode[1].Test,
           IN_Error_Level_1        := "DB009_Faults".Fault_State_Grp_1_M1,
           IN_SWU_OK               := "DB619_State_MPart".SWU[1].SWU_OK,
           IN_Release_Foamingcycle := "DB619_State_MPart".Cycle[1].Shotrelease,
           IN_ExternalRel_Foaming  := TRUE,
           IN_ToleranceOK_Foaming  := TRUE,
           IN_Foaming_Active       := "DB619_State_MPart".Cycle[1].ShotRuns,
           IO_Status               := "DB619_State_MPart".Mixinghead[1]
         );
   //-----
END_REGION

REGION Network 6: Opening of MH-valves
   //__________________________________________________________________
   // Valve mixinghead 01:
   //
         A     "DB619_State_MPart".Mixinghead[1].Mixingheadvalve."01";
         =     "DB123_MH_IO_Signals".MH[1].OUT.MH.V_MH;
   //__________________________________________________________________
   // Valve mixinghead 02:
   //
         A     "DB619_State_MPart".Mixinghead[1].Mixingheadvalve."02";
         =     "DB123_MH_IO_Signals".MH[2].OUT.MH.V_MH;
   //__________________________________________________________________
   // Valve mixinghead 03:
   //
         A     "DB619_State_MPart".Mixinghead[1].Mixingheadvalve."03";
         =     "DB123_MH_IO_Signals".MH[3].OUT.MH.V_MH;
   //__________________________________________________________________
   // Valve mixinghead 04:
   //
         A     "DB619_State_MPart".Mixinghead[1].Mixingheadvalve."04";
         =     "DB123_MH_IO_Signals".MH[4].OUT.MH.V_MH;
   //__________________________________________________________________
   // Valve mixinghead 05:
   //
         A     "DB619_State_MPart".Mixinghead[1].Mixingheadvalve."05";
         =     "DB123_MH_IO_Signals".MH[5].OUT.MH.V_MH;
   //__________________________________________________________________
   // Valve mixinghead 06:
   //
         A     "DB619_State_MPart".Mixinghead[1].Mixingheadvalve."06";
         =     "DB123_MH_IO_Signals".MH[6].OUT.MH.V_MH;
   //__________________________________________________________________
   // Valve mixinghead 07:
   //
         A     "DB619_State_MPart".Mixinghead[1].Mixingheadvalve."07";
         =     "DB123_MH_IO_Signals".MH[7].OUT.MH.V_MH;
   //__________________________________________________________________
   // Valve mixinghead 08:
   //
         A     "DB619_State_MPart".Mixinghead[1].Mixingheadvalve."08";
         =     "DB123_MH_IO_Signals".MH[8].OUT.MH.V_MH;
   //__________________________________________________________________
   // Valve mixinghead 08:
   //
         A     "DB619_State_MPart".Mixinghead[1].Mixingheadvalve."09";
         =     "DB123_MH_IO_Signals".MH[9].OUT.MH.V_MH;
   //__________________________________________________________________
   // Valve mixinghead 08:
   //
         A     "DB619_State_MPart".Mixinghead[1].Mixingheadvalve."10";
         =     "DB123_MH_IO_Signals".MH[10].OUT.MH.V_MH;
   //__________________________________________________________________
   //
END_REGION

REGION Network 7: Shotcounter
   //__________________________________________________________________
   // Shotcounter mixinghead 01:
   //
         A     "DB619_State_MPart".Mixinghead[1].Shotcounter."01";
         =     "DB123_MH_IO_Signals".MH[1].OUT.MH.H_Shotcounter_MH;
         JCN   countMH1end;
   //
         A     "DB619_State_MPart".Mixinghead[1].ImpCounterOn;
         JCN   countMH1end;
   //-----
         L     "DB_Zaehler_Anzeige".MH_Counter_Reset[1];
         L     1.0;
         +R;
         T     "DB_Zaehler_Anzeige".MH_Counter_Reset[1];
   //-----
         L     "DB_Zaehler_Anzeige".MH_Counter_NonReset[1];
         L     1.0;
         +R;
         T     "DB_Zaehler_Anzeige".MH_Counter_NonReset[1];
   //-----
         L     "DB_Zaehler_Schicht_aktuell".MH_Counter[1];
         L     1.0;
         +R;
         T     "DB_Zaehler_Schicht_aktuell".MH_Counter[1];
   //-----
   countMH1end:NOP   0;
   //__________________________________________________________________
   // Shotcounter mixinghead 02:
   //
         A     "DB619_State_MPart".Mixinghead[1].Shotcounter."02";
         =     "DB123_MH_IO_Signals".MH[2].OUT.MH.H_Shotcounter_MH;
         JCN   countMH2end;
   //
         A     "DB619_State_MPart".Mixinghead[1].ImpCounterOn;
         JCN   countMH2end;
   //-----
         L     "DB_Zaehler_Anzeige".MH_Counter_Reset[2];
         L     "DB619_State_MPart".Mixinghead[1].Countervalue;
         DTR;
         +R;
         T     "DB_Zaehler_Anzeige".MH_Counter_Reset[2];
   //-----
         L     "DB_Zaehler_Anzeige".MH_Counter_NonReset[2];
         L     "DB619_State_MPart".Mixinghead[1].Countervalue;
         DTR;
         +R;
         T     "DB_Zaehler_Anzeige".MH_Counter_NonReset[2];
   //-----
         L     "DB_Zaehler_Schicht_aktuell".MH_Counter[2];
         L     1.0;
         +R;
         T     "DB_Zaehler_Schicht_aktuell".MH_Counter[2];
   //-----
   countMH2end:NOP   0;
   //__________________________________________________________________
   // Shotcounter mixinghead 03:

         A     "DB619_State_MPart".Mixinghead[1].Shotcounter."03";
         =     "DB123_MH_IO_Signals".MH[3].OUT.MH.H_Shotcounter_MH;
         JCN   countMH3end;
   //
         A     "DB619_State_MPart".Mixinghead[1].ImpCounterOn;
         JCN   countMH3end;
   //-----
         L     "DB_Zaehler_Anzeige".MH_Counter_Reset[3];
         L     "DB619_State_MPart".Mixinghead[1].Countervalue;
         DTR;
         +R;
         T     "DB_Zaehler_Anzeige".MH_Counter_Reset[3];
   //-----
         L     "DB_Zaehler_Anzeige".MH_Counter_NonReset[3];
         L     "DB619_State_MPart".Mixinghead[1].Countervalue;
         DTR;
         +R;
         T     "DB_Zaehler_Anzeige".MH_Counter_NonReset[3];
   //-----
         L     "DB_Zaehler_Schicht_aktuell".MH_Counter[3];
         L     1.0;
         +R;
         T     "DB_Zaehler_Schicht_aktuell".MH_Counter[3];
   //-----
   countMH3end:NOP   0;
   //__________________________________________________________________
   // Shotcounter mixinghead 04:
   //
         A     "DB619_State_MPart".Mixinghead[1].Shotcounter."04";
         =     "DB123_MH_IO_Signals".MH[4].OUT.MH.H_Shotcounter_MH;
         JCN   countMH4end;
   //
         A     "DB619_State_MPart".Mixinghead[1].ImpCounterOn;
         JCN   countMH4end;
   //-----
         L     "DB_Zaehler_Anzeige".MH_Counter_Reset[4];
         L     "DB619_State_MPart".Mixinghead[1].Countervalue;
         DTR;
         +R;
         T     "DB_Zaehler_Anzeige".MH_Counter_Reset[4];
   //-----
         L     "DB_Zaehler_Anzeige".MH_Counter_NonReset[4];
         L     "DB619_State_MPart".Mixinghead[1].Countervalue;
         DTR;
         +R;
         T     "DB_Zaehler_Anzeige".MH_Counter_NonReset[4];
   //-----
         L     "DB_Zaehler_Schicht_aktuell".MH_Counter[4];
         L     1.0;
         +R;
         T     "DB_Zaehler_Schicht_aktuell".MH_Counter[4];
   //-----
   countMH4end:NOP   0;
   //__________________________________________________________________
   // Shotcounter mixinghead 05:
   //
         A     "DB619_State_MPart".Mixinghead[1].Shotcounter."05";
         =     "DB123_MH_IO_Signals".MH[5].OUT.MH.H_Shotcounter_MH;
         JCN   countMH5end;
   //
         A     "DB619_State_MPart".Mixinghead[1].ImpCounterOn;
         JCN   countMH5end;
   //-----
         L     "DB_Zaehler_Anzeige".MH_Counter_Reset[5];
         L     "DB619_State_MPart".Mixinghead[1].Countervalue;
         DTR;
         +R;
         T     "DB_Zaehler_Anzeige".MH_Counter_Reset[5];
   //-----
         L     "DB_Zaehler_Anzeige".MH_Counter_NonReset[5];
         L     "DB619_State_MPart".Mixinghead[1].Countervalue;
         DTR;
         +R;
         T     "DB_Zaehler_Anzeige".MH_Counter_NonReset[5];
   //-----
         L     "DB_Zaehler_Schicht_aktuell".MH_Counter[5];
         L     1.0;
         +R;
         T     "DB_Zaehler_Schicht_aktuell".MH_Counter[5];
   //-----
   countMH5end:NOP   0;
   //__________________________________________________________________
   // Shotcounter mixinghead 06:
   //
         A     "DB619_State_MPart".Mixinghead[1].Shotcounter."06";
         =     "DB123_MH_IO_Signals".MH[6].OUT.MH.H_Shotcounter_MH;
         JCN   countMH6end;
   //
         A     "DB619_State_MPart".Mixinghead[1].ImpCounterOn;
         JCN   countMH6end;
   //-----
         L     "DB_Zaehler_Anzeige".MH_Counter_Reset[6];
         L     "DB619_State_MPart".Mixinghead[1].Countervalue;
         DTR;
         +R;
         T     "DB_Zaehler_Anzeige".MH_Counter_Reset[6];
   //-----
         L     "DB_Zaehler_Anzeige".MH_Counter_NonReset[6];
         L     "DB619_State_MPart".Mixinghead[1].Countervalue;
         DTR;
         +R;
         T     "DB_Zaehler_Anzeige".MH_Counter_NonReset[6];
   //-----
         L     "DB_Zaehler_Schicht_aktuell".MH_Counter[6];
         L     1.0;
         +R;
         T     "DB_Zaehler_Schicht_aktuell".MH_Counter[6];
   //-----
   countMH6end:NOP   0;
   //__________________________________________________________________
   // Shotcounter mixinghead 07:
   //
         A     "DB619_State_MPart".Mixinghead[1].Shotcounter."07";
         =     "DB123_MH_IO_Signals".MH[7].OUT.MH.H_Shotcounter_MH;
         JCN   countMH7end;
   //
         A     "DB619_State_MPart".Mixinghead[1].ImpCounterOn;
         JCN   countMH7end;
   //-----
         L     "DB_Zaehler_Anzeige".MH_Counter_Reset[7];
         L     "DB619_State_MPart".Mixinghead[1].Countervalue;
         DTR;
         +R;
         T     "DB_Zaehler_Anzeige".MH_Counter_Reset[7];
   //-----
         L     "DB_Zaehler_Anzeige".MH_Counter_NonReset[7];
         L     "DB619_State_MPart".Mixinghead[1].Countervalue;
         DTR;
         +R;
         T     "DB_Zaehler_Anzeige".MH_Counter_NonReset[7];
   //-----
         L     "DB_Zaehler_Schicht_aktuell".MH_Counter[7];
         L     1.0;
         +R;
         T     "DB_Zaehler_Schicht_aktuell".MH_Counter[7];
   //-----
   countMH7end:NOP   0;